// TIA Portal project "PLC via Modbus to Arduino" (V17)

(* hardware
DEVICE "S7-1200 station_1"  S7-1200 Station
   slot 0: "Rack_0"  S7-1200 Rack  Rack  V1.0
   slot 1: "PLC_1"  CPU 1215C DC/DC/DC  6ES7 215-1AG40-0XB0  V4.4
   slot 101: "CM 1241 (RS422/485)_1"  6ES7 241-1CH32-0XB0  V2.2
DEVICE "HMI_1"  KTP700 Basic PN
   slot 0: "HMI_1"  KTP700 Basic PN  6AV2 123-2GB03-0AX0  17.0.0.0
   slot 1: "HMI_RT_1"  KTP700 Basic PN  6AV2 123-2GB03-0AX0  17.0.0.0
   slot 5: "HMI_1.IE_CP_1"  PROFINET Interface  17.0.0.0
      slot 1: "PROFINET Interface_1"  PROFINET Interface
         slot 1: "Port_1"  Port
*)

// ===== PLC "PLC_1"  CPU 1215C DC/DC/DC =====

VAR_GLOBAL   // PLC tag table "Default tag table"
   "System_Byte" AT %MB1 : Byte;
   "FirstScan" AT %M1.0 : Bool;
   "DiagStatusUpdate" AT %M1.1 : Bool;
   "AlwaysTRUE" AT %M1.2 : Bool;
   "AlwaysFALSE" AT %M1.3 : Bool;
   "Clock_Byte" AT %MB0 : Byte;
   "Clock_10Hz" AT %M0.0 : Bool;
   "Clock_5Hz" AT %M0.1 : Bool;
   "Clock_2.5Hz" AT %M0.2 : Bool;
   "Clock_2Hz" AT %M0.3 : Bool;
   "Clock_1.25Hz" AT %M0.4 : Bool;
   "Clock_1Hz" AT %M0.5 : Bool;
   "Clock_0.625Hz" AT %M0.6 : Bool;
   "Clock_0.5Hz" AT %M0.7 : Bool;
   "Run_Cycle" AT %M10.0 : Bool;
   "Request_Temperature" AT %M10.1 : Bool;
   "Request_Humidity" AT %M10.2 : Bool;
   "Read_Temperature" AT %MW100 : Int;
   "Read_Humidity" AT %MW102 : Int;
   "Cycle_Case" AT %MW104 : Int;
   "Pulse_Time" AT %MD200 : Time;
   "Read_Delay" AT %MD204 : Time;
END_VAR

// folder: System blocks/Program resources

DATA_BLOCK "IEC_Timer_0_DB"   // DB3
{ S7_Optimized_Access := 'TRUE' }
AUTHOR : Simatic
FAMILY : IEC
NAME : IEC_TMR
VERSION : 1.0
// stored: InstanceOfName IEC_TIMER
"IEC_TIMER"
BEGIN
END_DATA_BLOCK

DATA_BLOCK "IEC_Timer_0_DB_1"   // DB4
{ S7_Optimized_Access := 'TRUE' }
AUTHOR : Simatic
FAMILY : IEC
NAME : IEC_TMR
VERSION : 1.0
// stored: InstanceOfName IEC_TIMER
"IEC_TIMER"
BEGIN
END_DATA_BLOCK

DATA_BLOCK "IEC_Timer_0_DB_2"   // DB5
{ S7_Optimized_Access := 'TRUE' }
AUTHOR : Simatic
FAMILY : IEC
NAME : IEC_TMR
VERSION : 1.0
// stored: InstanceOfName IEC_TIMER
"IEC_TIMER"
BEGIN
END_DATA_BLOCK

DATA_BLOCK "IEC_Timer_0_DB_3"   // DB6
{ S7_Optimized_Access := 'TRUE' }
AUTHOR : Simatic
FAMILY : IEC
NAME : IEC_TMR
VERSION : 1.0
// stored: InstanceOfName IEC_TIMER
"IEC_TIMER"
BEGIN
END_DATA_BLOCK

// folder: (top level)

FUNCTION "RS485_Comms" : Void   // FC1, LAD
{ S7_Optimized_Access := 'TRUE' }
VERSION : 0.1
   VAR_TEMP   // added for the SCL form of the ladder/FBD networks
      _w1 : Bool;
   END_VAR
BEGIN

REGION Network 1
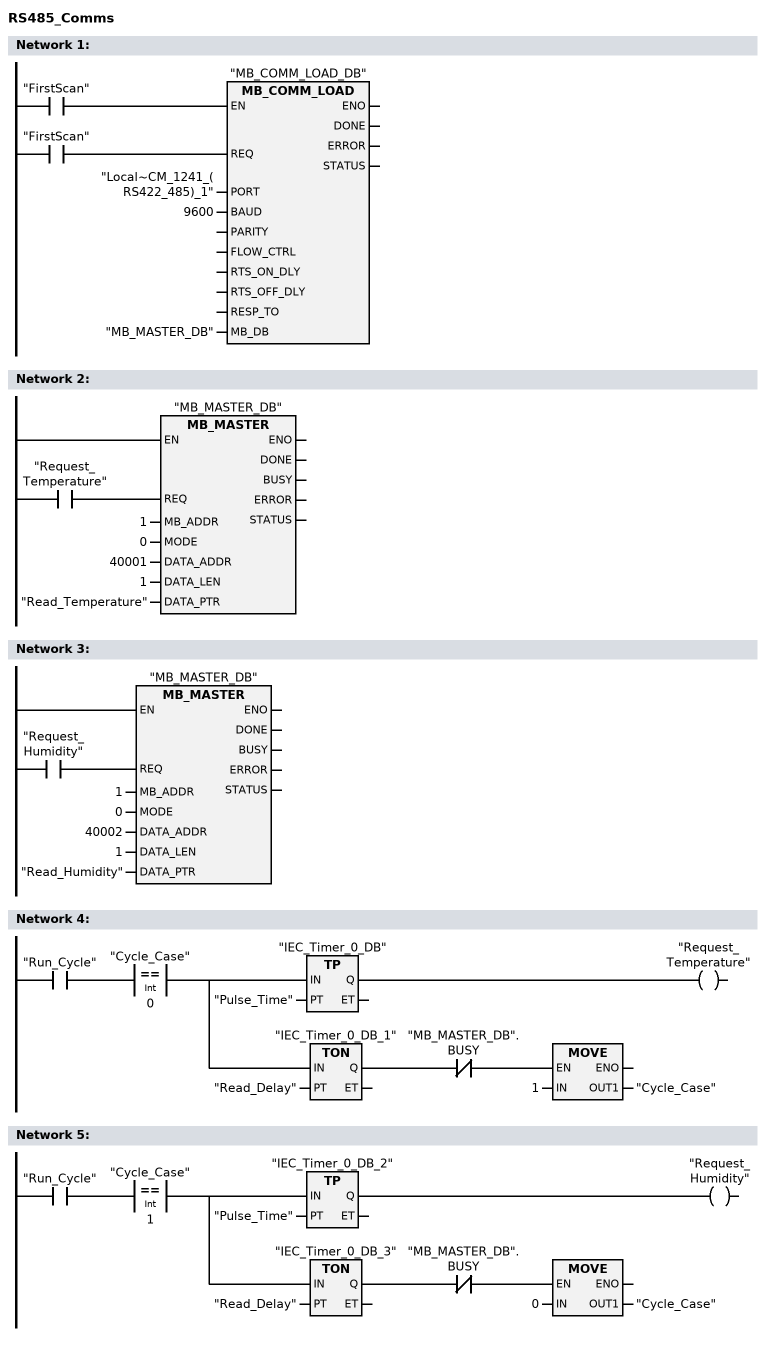
   IF "FirstScan" THEN
       "MB_COMM_LOAD_DB"(REQ := "FirstScan",   // MB_COMM_LOAD
                         PORT := "Local~CM_1241_(RS422_485)_1",
                         BAUD := 9600,
                         MB_DB := "MB_MASTER_DB");
   END_IF;
END_REGION

REGION Network 2
   "MB_MASTER_DB"(REQ := "Request_Temperature",   // MB_MASTER
                  MB_ADDR := 1,
                  MODE := 0,
                  DATA_ADDR := 40001,
                  DATA_LEN := 1,
                  DATA_PTR := "Read_Temperature");
END_REGION

REGION Network 3
   "MB_MASTER_DB"(REQ := "Request_Humidity",   // MB_MASTER
                  MB_ADDR := 1,
                  MODE := 0,
                  DATA_ADDR := 40002,
                  DATA_LEN := 1,
                  DATA_PTR := "Read_Humidity");
END_REGION

REGION Network 4
   #_w1 := "Run_Cycle" AND ("Cycle_Case" = 0);
   "IEC_Timer_0_DB".TP(IN := #_w1, PT := "Pulse_Time");
   "Request_Temperature" := "IEC_Timer_0_DB".Q;
   "IEC_Timer_0_DB_1".TON(IN := #_w1, PT := "Read_Delay");
   IF "IEC_Timer_0_DB_1".Q AND NOT "MB_MASTER_DB".BUSY THEN "Cycle_Case" := 1; END_IF;
END_REGION

REGION Network 5
   #_w1 := "Run_Cycle" AND ("Cycle_Case" = 1);
   "IEC_Timer_0_DB_2".TP(IN := #_w1, PT := "Pulse_Time");
   "Request_Humidity" := "IEC_Timer_0_DB_2".Q;
   "IEC_Timer_0_DB_3".TON(IN := #_w1, PT := "Read_Delay");
   IF "IEC_Timer_0_DB_3".Q AND NOT "MB_MASTER_DB".BUSY THEN "Cycle_Case" := 0; END_IF;
END_REGION
END_FUNCTION

ORGANIZATION_BLOCK "Main"   // OB1, LAD, ProgramCycle
TITLE = "Main Program Sweep (Cycle)"
{ S7_Optimized_Access := 'TRUE' }
VERSION : 0.1
   VAR_INPUT
      Initial_Call : Bool;   // Initial call of this OB
      Remanence : Bool;   // =True, if remanent data are available
   END_VAR
BEGIN

REGION Network 1
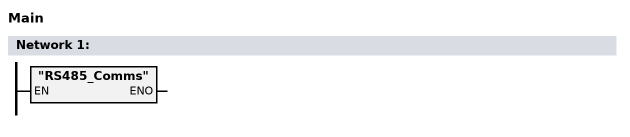
   RUNG wire#powerrail
      "RS485_Comms"()
   END_RUNG
   // the same network as SCL:
   "RS485_Comms"();
END_REGION
END_ORGANIZATION_BLOCK

(* ===== HMI "HMI_RT_1" =====
system functions are stored by id; their names below are inferred from use
connection "HMI_Connection_1": ETHERNET, SMART_S7_1200_OMS

HMI tags "Default tag table"
   "Tag_ScreenNumber" : UInt, internal
   "readTemperature" : Int = PLC Read_Temperature AT %MW100, 100 ms
   "readHumidity" : Int = PLC Read_Humidity AT %MW102, 100 ms
   "setPulseTime" : Time = PLC Pulse_Time AT %MD200, 1 s
   "setReadDelay" : Time = PLC Read_Delay AT %MD204, 1 s
   "startCycle" : Bool = PLC Run_Cycle AT %M10.0, 1 s

Template "Template_1" 800x480
   Button "Exit" at 714,429 size 71x50; TextOff 'Exit'; PictureOff "ExitRuntime_KTP700_Basic_PN_TR"; PictureOn "ExitRuntime_KTP700_Basic_PN_TR"
      on Release: StopRuntime(0)
   Button "Template_Button" at 614,429 size 71x50; TextOff 'Text'
   Button "Template_Button_1" at 514,429 size 71x50; TextOff 'Text'
   Button "Template_Button_2" at 414,429 size 71x50; TextOff 'Text'
   Button "Template_Button_3" at 314,429 size 71x50; TextOff 'Text'
   Button "Template_Button_4" at 214,429 size 71x50; TextOff 'Text'
   Button "Template_Button_5" at 114,429 size 71x50; TextOff 'Text'
   Button "Start screen" at 14,429 size 71x50; TextOff 'Start screen'; PictureOff "NavigateHome_KTP700_Basic_PN_TR"; PictureOn "NavigateHome_KTP700_Basic_PN_TR"
      on Release: ActivateScreen("Root screen", 0)
   SymbolicIOField "Symbolic_IO_Field_Screen" at 93,9 size 600x33; TextOff '0'; TextOn '1'; TextList "TextList_ScreenNames"
      ProcessValue <- "Tag_ScreenNumber"
      on Change: ActivateScreenByNumber("Tag_ScreenNumber", 0)
   DateTimeField "HmiScreenItemData" at 695,25 size 105x25
   DateTimeField "HmiScreenItemData_1" at 695,0 size 105x25
   GraphicView "Logo" at 0,0 size 91x51; Picture "Logo of HMI_1"

screen "Root screen" 800x480
   on GenerateScreen: SetTag("Tag_ScreenNumber", 1)
   TextField "Text field_1" at 167,126 size 118x23; Text 'Temperature:'
   IOField "I/O field_1" at 287,123 size 96x32; FormatPattern 9999
      ProcessValue <- "readTemperature"
   TextField "Text field_2" at 167,174 size 84x23; Text 'Humidity:'
   IOField "I/O field_2" at 287,171 size 96x32; FormatPattern 9999
      ProcessValue <- "readHumidity"
   TextField "Text field_3" at 403,126 size 101x23; Text 'Pulse Time:'
   IOField "I/O field_3" at 523,123 size 96x32; FormatPattern 9999
      ProcessValue <- "setPulseTime"
   TextField "Text field_4" at 403,174 size 104x23; Text 'Read Delay:'
   IOField "I/O field_4" at 523,171 size 96x32; FormatPattern 9999
      ProcessValue <- "setReadDelay"
   Switch "Switch_1" at 241,246 size 324x32; CaptionText 'Switch'; TextOff 'Not Running'; TextOn 'Running'
      ProcessValue <- "startCycle"
*)